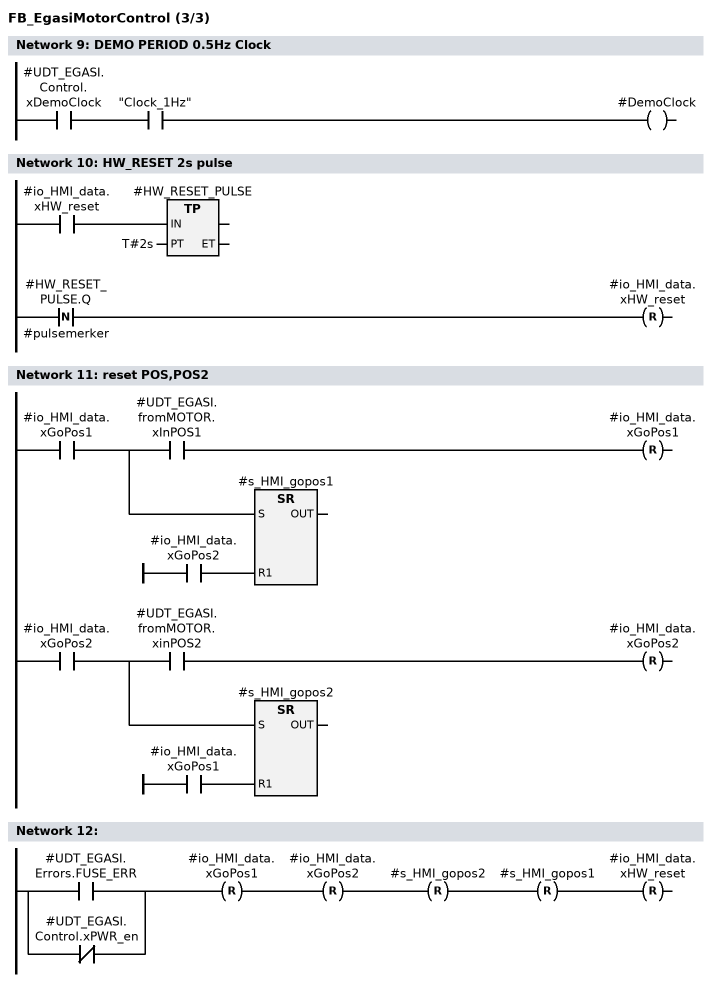
   RUNG wire#powerrail
      Contact( #UDT_EGASI.Control.xDemoClock )
      Contact( "Clock_1Hz" )
      Coil( #DemoClock )
   END_RUNG
   // the same network as SCL:
   #DemoClock := #UDT_EGASI.Control.xDemoClock AND "Clock_1Hz";
END_REGION

REGION Network 10: HW_RESET 2s pulse
   #HW_RESET_PULSE(IN := #io_HMI_data.xHW_reset, PT := T#2s);   // TP
   #_w1 := NOT #HW_RESET_PULSE.Q AND #pulsemerker;   // falling edge of #HW_RESET_PULSE.Q
   #pulsemerker := #HW_RESET_PULSE.Q;
   IF #_w1 THEN #io_HMI_data.xHW_reset := FALSE; END_IF;
END_REGION

REGION Network 11: reset POS,POS2
   RUNG wire#powerrail
      Contact( #io_HMI_data.xGoPos1 )
      wire#w1
      Contact( #UDT_EGASI.fromMOTOR.xInPOS1 )
      R_Coil( #io_HMI_data.xGoPos1 )
   END_RUNG
   RUNG wire#w1
      S_SR(operand := #s_HMI_gopos1, r1 := wire#w2)
   END_RUNG
   RUNG wire#powerrail
      Contact( #io_HMI_data.xGoPos2 )
   END_RUNG wire#w2
   RUNG wire#powerrail
      Contact( #io_HMI_data.xGoPos2 )
      wire#w3
      Contact( #UDT_EGASI.fromMOTOR.xinPOS2 )
      R_Coil( #io_HMI_data.xGoPos2 )
   END_RUNG
   RUNG wire#w3
      S_SR(operand := #s_HMI_gopos2, r1 := wire#w4)
   END_RUNG
   RUNG wire#powerrail
      Contact( #io_HMI_data.xGoPos1 )
   END_RUNG wire#w4
   // the same network as SCL:
   #_w1 := #io_HMI_data.xGoPos1;
   IF #io_HMI_data.xGoPos1 AND #UDT_EGASI.fromMOTOR.xInPOS1 THEN #io_HMI_data.xGoPos1 := FALSE; END_IF;
   IF #_w1 THEN
       #s_HMI_gopos1 := TRUE;   // SR flip-flop
   END_IF;
   IF #io_HMI_data.xGoPos2 THEN #s_HMI_gopos1 := FALSE; END_IF;
   #_w2 := #io_HMI_data.xGoPos2;
   IF #io_HMI_data.xGoPos2 AND #UDT_EGASI.fromMOTOR.xinPOS2 THEN #io_HMI_data.xGoPos2 := FALSE; END_IF;
   IF #_w2 THEN
       #s_HMI_gopos2 := TRUE;   // SR flip-flop
   END_IF;
   IF #io_HMI_data.xGoPos1 THEN #s_HMI_gopos2 := FALSE; END_IF;
END_REGION

REGION Network 12
   RUNG wire#powerrail
      Contact( #UDT_EGASI.Errors.FUSE_ERR )
      wire#w1
      R_Coil( #io_HMI_data.xGoPos1 )
      R_Coil( #io_HMI_data.xGoPos2 )
      R_Coil( #s_HMI_gopos2 )
      R_Coil( #s_HMI_gopos1 )
      R_Coil( #io_HMI_data.xHW_reset )
   END_RUNG
   RUNG wire#powerrail
      I_Contact( #UDT_EGASI.Control.xPWR_en )
   END_RUNG wire#w1
   // the same network as SCL:
   IF #UDT_EGASI.Errors.FUSE_ERR OR NOT #UDT_EGASI.Control.xPWR_en THEN
       #io_HMI_data.xGoPos1 := FALSE;
       #io_HMI_data.xGoPos2 := FALSE;
       #s_HMI_gopos2 := FALSE;
       #s_HMI_gopos1 := FALSE;
       #io_HMI_data.xHW_reset := FALSE;
   END_IF;
END_REGION

REGION Network 13 (SCL)
   #q_rScaledTemperature := ((#i_wRawTempValue/32767.0) * 10.0)/0.04;
   #UDT_EGASI.fromMOTOR.wRawTempValue := #i_wRawTempValue;
   #UDT_EGASI.fromMOTOR.rScaledTempValue := #q_rScaledTemperature;
END_REGION
END_FUNCTION_BLOCK

FUNCTION_BLOCK "FB_Convert16bitToTemperature"   // FB17, LAD
{ S7_Optimized_Access := 'TRUE' }
VERSION : 0.1
   VAR_INPUT
      i_wRawValue : Word;
   END_VAR
   VAR_OUTPUT
      q_uiScaledTemperature : Real;
   END_VAR
BEGIN

REGION Network 2 (SCL)
   #q_uiScaledTemperature := #i_wRawValue/32767.0 * 0.04;
END_REGION
END_FUNCTION_BLOCK

FUNCTION_BLOCK "FB_CYLINDER_CONTROL"   // FB18, LAD
{ S7_Optimized_Access := 'TRUE' }
VERSION : 0.1
   VAR_INPUT
      i_xTrigger : Bool;
      i_udMAXDontProduceFeedCounter : UDInt;
   END_VAR
   VAR_OUTPUT
      q_xM1Output : Bool;
      q_xM2Output : Bool;
      q_xM3Output : Bool;
      q_xM4Output : Bool;
      q_xM5Output : Bool;
   END_VAR
   VAR_IN_OUT
      io_CylinderData : "RRI_izdelki";
      io_LastCylinderData : "RRI_izdelki";
      io_ReceptToMake : "RRI_izdelki";
      io_xChangingPart : Bool;
      io_xuiChangePartCounter : UDInt;
      io_iTrenutniPomik : Int;
      PartNumberForProduction : String;
      LastPartForProduction : String;
   END_VAR
   VAR RETAIN
      markers : Array[0..1] of Bool;
      ChangePartStepCounter : Int;
      iLastPartStVrst : Int;
      iLastPartStCelic : Int;
   END_VAR
   VAR_TEMP   // added for the SCL form of the ladder/FBD networks
      _w1 : Bool;
   END_VAR
BEGIN

REGION Network 1: Povečaj števec za trenutni števec
   // pocečaj trneutni pomik
   // povečaj pomik, če je
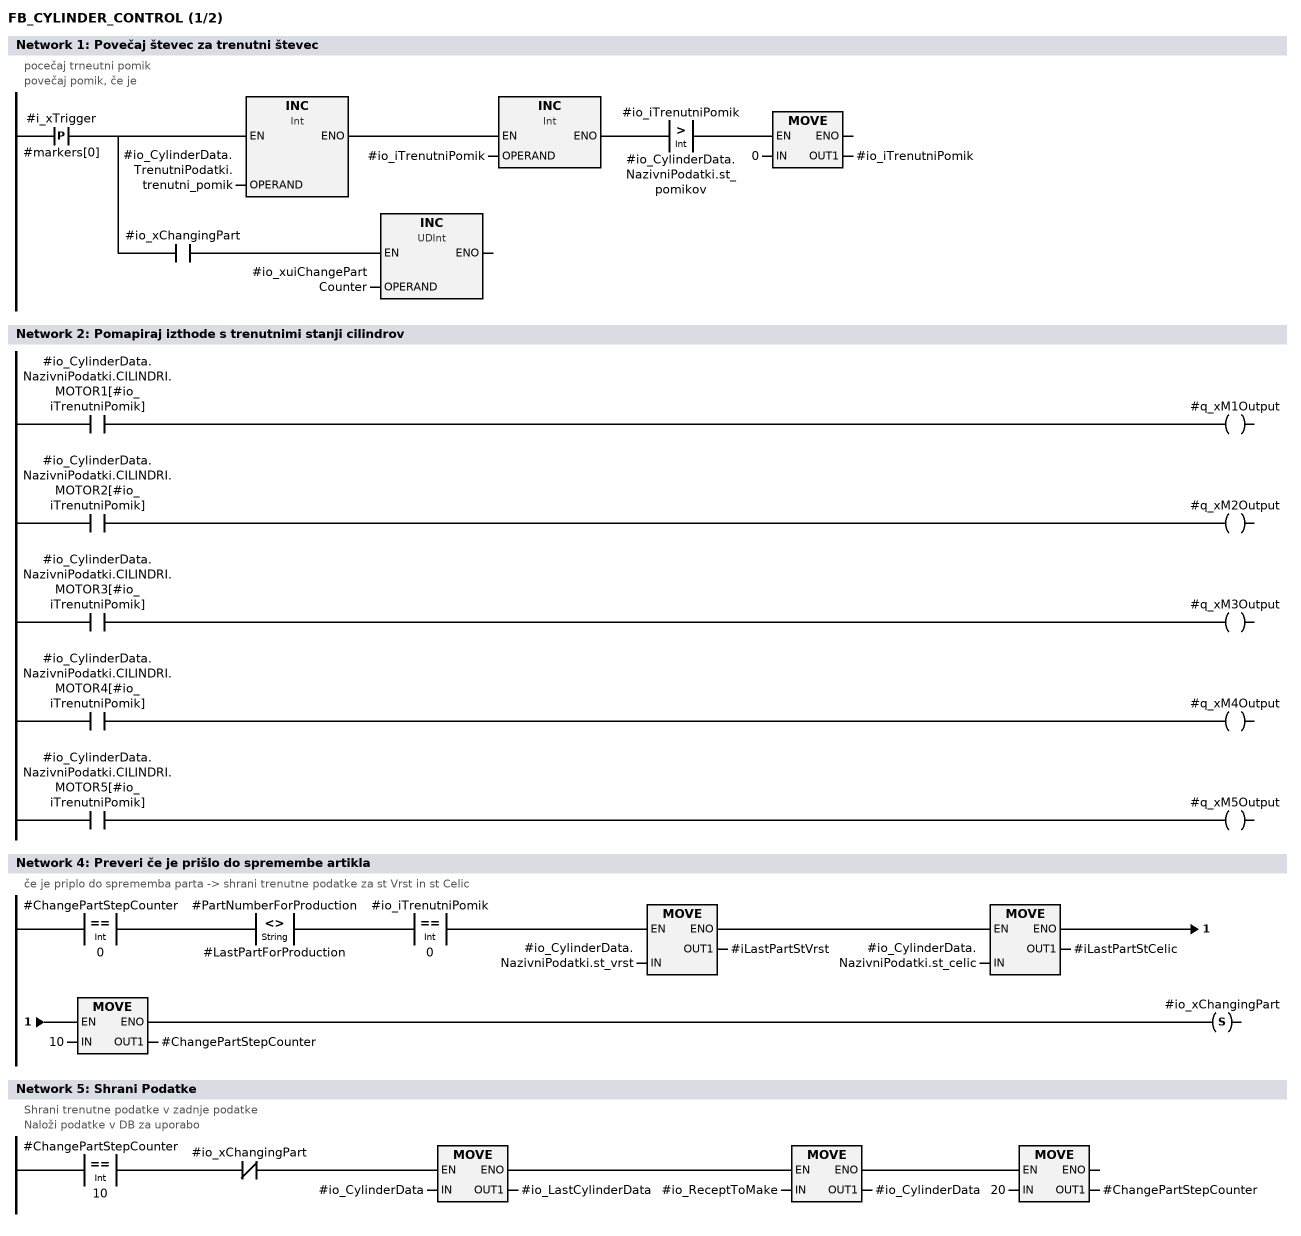
   RUNG wire#powerrail
      P_Contact(operand := #i_xTrigger, bit := #markers[0])
      wire#w1
      { S7_Templates := "DestType := Int" } Inc( #io_CylinderData.TrenutniPodatki.trenutni_pomik )
      { S7_Templates := "DestType := Int" } Inc( #io_iTrenutniPomik )
      { S7_Templates := "SrcType := Int" } GT_Contact(in1 := #io_iTrenutniPomik, in2 := #io_CylinderData.NazivniPodatki.st_pomikov)
      Move(in := 0, out1 => #io_iTrenutniPomik)
   END_RUNG
   RUNG wire#w1
      Contact( #io_xChangingPart )
      { S7_Templates := "DestType := UDInt" } Inc( #io_xuiChangePartCounter )
   END_RUNG
   // the same network as SCL:
   #_w1 := #i_xTrigger AND NOT #markers[0];   // rising edge of #i_xTrigger
   #markers[0] := #i_xTrigger;
   IF #_w1 THEN
       #io_CylinderData.TrenutniPodatki.trenutni_pomik := #io_CylinderData.TrenutniPodatki.trenutni_pomik + 1;
       #io_iTrenutniPomik := #io_iTrenutniPomik + 1;
   END_IF;
   IF #_w1 AND (#io_iTrenutniPomik > #io_CylinderData.NazivniPodatki.st_pomikov) THEN
       #io_iTrenutniPomik := 0;
   END_IF;
   IF #_w1 AND #io_xChangingPart THEN #io_xuiChangePartCounter := #io_xuiChangePartCounter + 1; END_IF;
END_REGION

REGION Network 2: Pomapiraj izthode s trenutnimi stanji cilindrov
   RUNG wire#powerrail
      Contact( #io_CylinderData.NazivniPodatki.CILINDRI.MOTOR1[#io_iTrenutniPomik] )
      Coil( #q_xM1Output )
   END_RUNG
   RUNG wire#powerrail
      Contact( #io_CylinderData.NazivniPodatki.CILINDRI.MOTOR2[#io_iTrenutniPomik] )
      Coil( #q_xM2Output )
   END_RUNG
   RUNG wire#powerrail
      Contact( #io_CylinderData.NazivniPodatki.CILINDRI.MOTOR3[#io_iTrenutniPomik] )
      Coil( #q_xM3Output )
   END_RUNG
   RUNG wire#powerrail
      Contact( #io_CylinderData.NazivniPodatki.CILINDRI.MOTOR4[#io_iTrenutniPomik] )
      Coil( #q_xM4Output )
   END_RUNG
   RUNG wire#powerrail
      Contact( #io_CylinderData.NazivniPodatki.CILINDRI.MOTOR5[#io_iTrenutniPomik] )
      Coil( #q_xM5Output )
   END_RUNG
   // the same network as SCL:
   #q_xM1Output := #io_CylinderData.NazivniPodatki.CILINDRI.MOTOR1[#io_iTrenutniPomik];
   #q_xM2Output := #io_CylinderData.NazivniPodatki.CILINDRI.MOTOR2[#io_iTrenutniPomik];
   #q_xM3Output := #io_CylinderData.NazivniPodatki.CILINDRI.MOTOR3[#io_iTrenutniPomik];
   #q_xM4Output := #io_CylinderData.NazivniPodatki.CILINDRI.MOTOR4[#io_iTrenutniPomik];
   #q_xM5Output := #io_CylinderData.NazivniPodatki.CILINDRI.MOTOR5[#io_iTrenutniPomik];
END_REGION

REGION Network 4: Preveri če je prišlo do spremembe artikla
   // če je priplo do sprememba parta -> shrani trenutne podatke za st Vrst in st Celic
   RUNG wire#powerrail
      { S7_Templates := "SrcType := Int" } EQ_Contact(in1 := #ChangePartStepCounter, in2 := 0)
      { S7_Templates := "SrcType := String" } NE_Contact(in1 := #PartNumberForProduction, in2 := #LastPartForProduction)
      { S7_Templates := "SrcType := Int" } EQ_Contact(in1 := #io_iTrenutniPomik, in2 := 0)
      Move(in := #io_CylinderData.NazivniPodatki.st_vrst, out1 => #iLastPartStVrst)
      Move(in := #io_CylinderData.NazivniPodatki.st_celic, out1 => #iLastPartStCelic)
      Move(in := 10, out1 => #ChangePartStepCounter)
      S_Coil( #io_xChangingPart )
   END_RUNG
   // the same network as SCL:
   IF (#ChangePartStepCounter = 0) AND (#PartNumberForProduction <> #LastPartForProduction) AND (#io_iTrenutniPomik = 0) THEN
       #iLastPartStVrst := #io_CylinderData.NazivniPodatki.st_vrst;
       #iLastPartStCelic := #io_CylinderData.NazivniPodatki.st_celic;
   END_IF;
   #_w1 := (#ChangePartStepCounter = 0) AND (#PartNumberForProduction <> #LastPartForProduction) AND (#io_iTrenutniPomik = 0);
   IF #_w1 THEN
       #ChangePartStepCounter := 10;
       #io_xChangingPart := TRUE;
   END_IF;
END_REGION

REGION Network 5: Shrani Podatke
   // Shrani trenutne podatke v zadnje podatke
   // Naloži podatke v DB za uporabo
   RUNG wire#powerrail
      { S7_Templates := "SrcType := Int" } EQ_Contact(in1 := #ChangePartStepCounter, in2 := 10)
      I_Contact( #io_xChangingPart )
      Move(in := #io_CylinderData, out1 => #io_LastCylinderData)
      Move(in := #io_ReceptToMake, out1 => #io_CylinderData)
      Move(in := 20, out1 => #ChangePartStepCounter)
   END_RUNG
   // the same network as SCL:
   IF (#ChangePartStepCounter = 10) AND NOT #io_xChangingPart THEN
       #io_LastCylinderData := #io_CylinderData;
       #io_CylinderData := #io_ReceptToMake;
       #ChangePartStepCounter := 20;
   END_IF;
END_REGION

REGION Network 6
   // Shrani partnumber
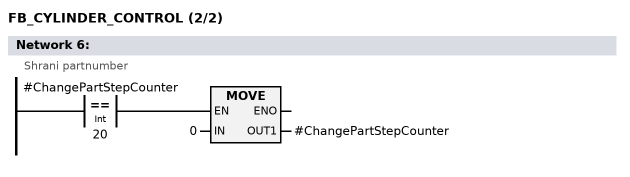
   RUNG wire#powerrail
      { S7_Templates := "SrcType := Int" } EQ_Contact(in1 := #ChangePartStepCounter, in2 := 20)
      Move(in := 0, out1 => #ChangePartStepCounter)
   END_RUNG
   // the same network as SCL:
   IF #ChangePartStepCounter = 20 THEN #ChangePartStepCounter := 0; END_IF;
END_REGION
END_FUNCTION_BLOCK

FUNCTION "FC_INPUT" : Void   // FC1, LAD
{ S7_Optimized_Access := 'TRUE' }
VERSION : 0.1
BEGIN

REGION Network 1: PLC input mapping
   // AKD1 - fault relay - open if error
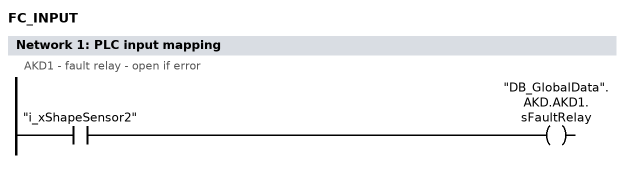
   RUNG wire#powerrail
      Contact( "i_xShapeSensor2" )
      Coil( "DB_GlobalData".AKD.AKD1.sFaultRelay )
   END_RUNG
   // the same network as SCL:
   "DB_GlobalData".AKD.AKD1.sFaultRelay := "i_xShapeSensor2";
END_REGION
END_FUNCTION

FUNCTION "FC_OUTPUT" : Void   // FC2, LAD
{ S7_Optimized_Access := 'TRUE' }
VERSION : 0.1
BEGIN

REGION Network 1: Communication mapping for NodeRed data and DATAFORCOMUNICATIONDB
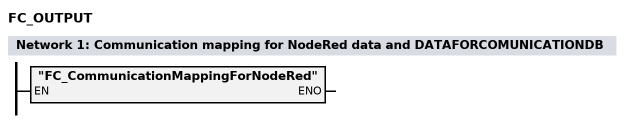
   RUNG wire#powerrail
      "FC_CommunicationMappingForNodeRed"()
   END_RUNG
   // the same network as SCL:
   "FC_CommunicationMappingForNodeRed"();
END_REGION
END_FUNCTION

FUNCTION "FC_LOGIC" : Void   // FC3, LAD
{ S7_Optimized_Access := 'TRUE' }
VERSION : 0.1
BEGIN

REGION Network 1: Convert ThermocuplerData
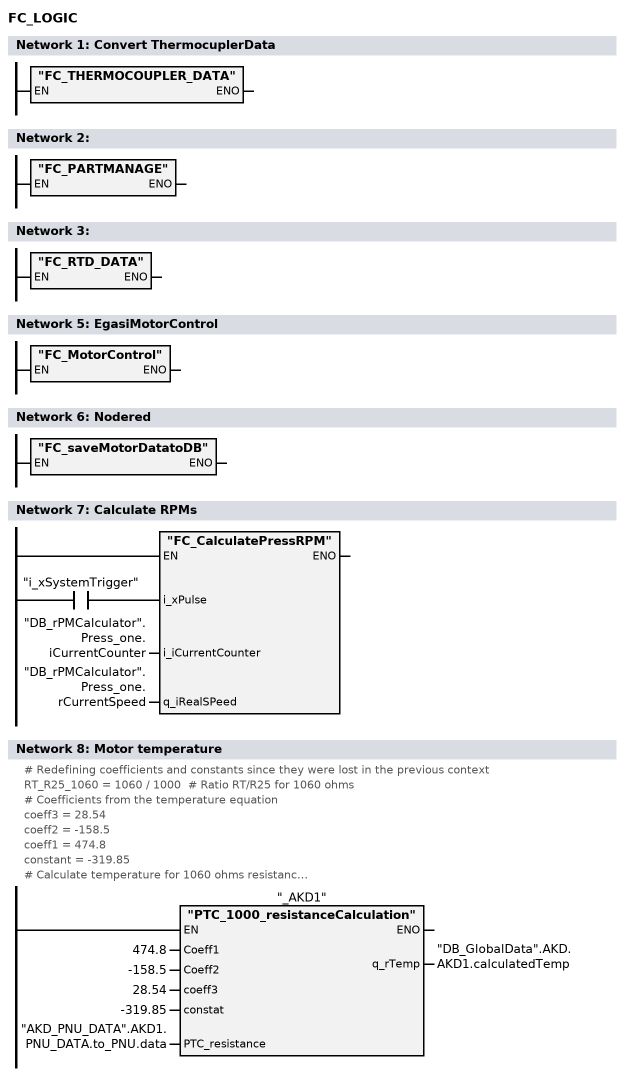
   RUNG wire#powerrail
      "FC_THERMOCOUPLER_DATA"()
   END_RUNG
   // the same network as SCL:
   "FC_THERMOCOUPLER_DATA"();
END_REGION

REGION Network 2
   RUNG wire#powerrail
      "FC_PARTMANAGE"()
   END_RUNG
   // the same network as SCL:
   "FC_PARTMANAGE"();
END_REGION

REGION Network 3
   RUNG wire#powerrail
      "FC_RTD_DATA"()
   END_RUNG
   // the same network as SCL:
   "FC_RTD_DATA"();
END_REGION

REGION Network 4: Kollmorgen Settings
END_REGION

REGION Network 5: EgasiMotorControl
   RUNG wire#powerrail
      "FC_MotorControl"()
   END_RUNG
   // the same network as SCL:
   "FC_MotorControl"();
END_REGION

REGION Network 6: Nodered
   RUNG wire#powerrail
      "FC_saveMotorDatatoDB"()
   END_RUNG
   // the same network as SCL:
   "FC_saveMotorDatatoDB"();
END_REGION

REGION Network 7: Calculate RPMs
   RUNG wire#powerrail
      "FC_CalculatePressRPM"(i_xPulse := wire#w1, i_iCurrentCounter := "DB_rPMCalculator".Press_one.iCurrentCounter, q_iRealSPeed := "DB_rPMCalculator".Press_one.rCurrentSpeed)
   END_RUNG
   RUNG wire#powerrail
      Contact( "i_xSystemTrigger" )
   END_RUNG wire#w1
   // the same network as SCL:
   "FC_CalculatePressRPM"(i_xPulse := "i_xSystemTrigger",
                          i_iCurrentCounter := "DB_rPMCalculator".Press_one.iCurrentCounter,
                          q_iRealSPeed := "DB_rPMCalculator".Press_one.rCurrentSpeed);
END_REGION

REGION Network 8: Motor temperature
   // # Redefining coefficients and constants since they were lost in the previous context
   // RT_R25_1060 = 1060 / 1000  # Ratio RT/R25 for 1060 ohms
   // 
   // # Coefficients from the temperature equation
   // coeff3 = 28.54
   // coeff2 = -158.5
   // coeff1 = 474.8
   // constant = -319.85
   // 
   // # Calculate temperature for 1060 ohms resistance
   // temperature_1060 = (coeff3 * RT_R25_1060**3) + (coeff2 * RT_R25_1060**2) + (coeff1 * RT_R25_1060) + constant
   RUNG wire#powerrail
      "_AKD1"(Coeff1 := 474.8, Coeff2 := -158.5, coeff3 := 28.54, constat := -319.85, PTC_resistance := "AKD_PNU_DATA".AKD1.PNU_DATA.to_PNU.data, q_rTemp => "DB_GlobalData".AKD.AKD1.calculatedTemp)
   END_RUNG
   // the same network as SCL:
   "_AKD1"(Coeff1 := 474.8,   // "PTC_1000_resistanceCalculation"
           Coeff2 := -158.5,
           coeff3 := 28.54,
           constat := -319.85,
           PTC_resistance := "AKD_PNU_DATA".AKD1.PNU_DATA.to_PNU.data,
           q_rTemp => "DB_GlobalData".AKD.AKD1.calculatedTemp);
END_REGION
END_FUNCTION

FUNCTION "FC_THERMOCOUPLER_DATA" : Void   // FC4, LAD
{ S7_Optimized_Access := 'TRUE' }
VERSION : 0.1
BEGIN

REGION Network 1: Temeprature conversion - from Input to GlobalDataBLock
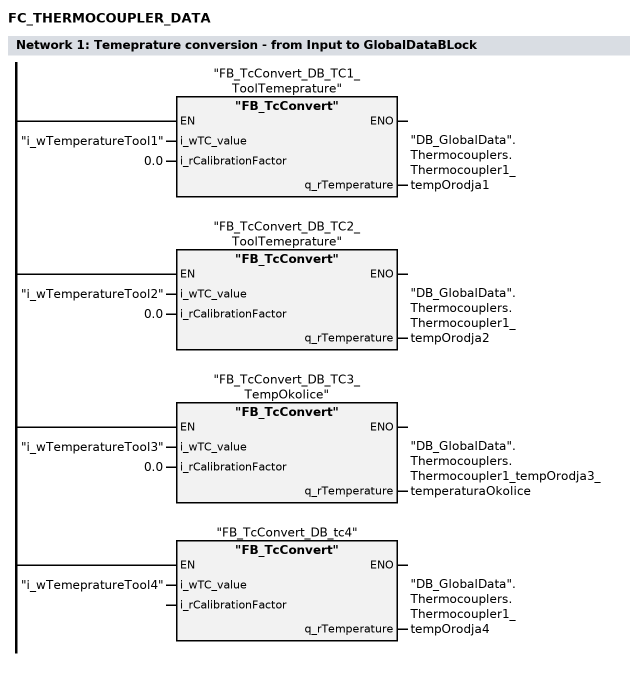
   RUNG wire#powerrail
      "FB_TcConvert_DB_TC1_ToolTemeprature"(i_wTC_value := "i_wTemperatureTool1", i_rCalibrationFactor := 0.0, q_rTemperature => "DB_GlobalData".Thermocouplers.Thermocoupler1_tempOrodja1)
   END_RUNG
   RUNG wire#powerrail
      "FB_TcConvert_DB_TC2_ToolTemeprature"(i_wTC_value := "i_wTemperatureTool2", i_rCalibrationFactor := 0.0, q_rTemperature => "DB_GlobalData".Thermocouplers.Thermocoupler1_tempOrodja2)
   END_RUNG
   RUNG wire#powerrail
      "FB_TcConvert_DB_TC3_TempOkolice"(i_wTC_value := "i_wTemperatureTool3", i_rCalibrationFactor := 0.0, q_rTemperature => "DB_GlobalData".Thermocouplers.Thermocoupler1_tempOrodja3_temperaturaOkolice)
   END_RUNG
   RUNG wire#powerrail
      "FB_TcConvert_DB_tc4"(i_wTC_value := "i_wTemepratureTool4", i_rCalibrationFactor :=, q_rTemperature => "DB_GlobalData".Thermocouplers.Thermocoupler1_tempOrodja4)
   END_RUNG
   // the same network as SCL:
   "FB_TcConvert_DB_TC1_ToolTemeprature"(i_wTC_value := "i_wTemperatureTool1",   // "FB_TcConvert"
                           i_rCalibrationFactor := 0.0,
                           q_rTemperature => "DB_GlobalData".Thermocouplers.Thermocoupler1_tempOrodja1);
   "FB_TcConvert_DB_TC2_ToolTemeprature"(i_wTC_value := "i_wTemperatureTool2",   // "FB_TcConvert"
                           i_rCalibrationFactor := 0.0,
                           q_rTemperature => "DB_GlobalData".Thermocouplers.Thermocoupler1_tempOrodja2);
   "FB_TcConvert_DB_TC3_TempOkolice"(i_wTC_value := "i_wTemperatureTool3",   // "FB_TcConvert"
                           i_rCalibrationFactor := 0.0,
                           q_rTemperature => "DB_GlobalData".Thermocouplers.Thermocoupler1_tempOrodja3_temperaturaOkolice);
   "FB_TcConvert_DB_tc4"(i_wTC_value := "i_wTemepratureTool4",   // "FB_TcConvert"
                         q_rTemperature => "DB_GlobalData".Thermocouplers.Thermocoupler1_tempOrodja4);
END_REGION
END_FUNCTION

FUNCTION "FC_CommunicationMappingForNodeRed" : Void   // FC5, LAD
{ S7_Optimized_Access := 'TRUE' }
VERSION : 0.1
   VAR_TEMP   // added for the SCL form of the ladder/FBD networks
      _w1 : Bool;
   END_VAR
BEGIN

REGION Network 1: Move data from GlobalData to DB for NodeRedCommunication
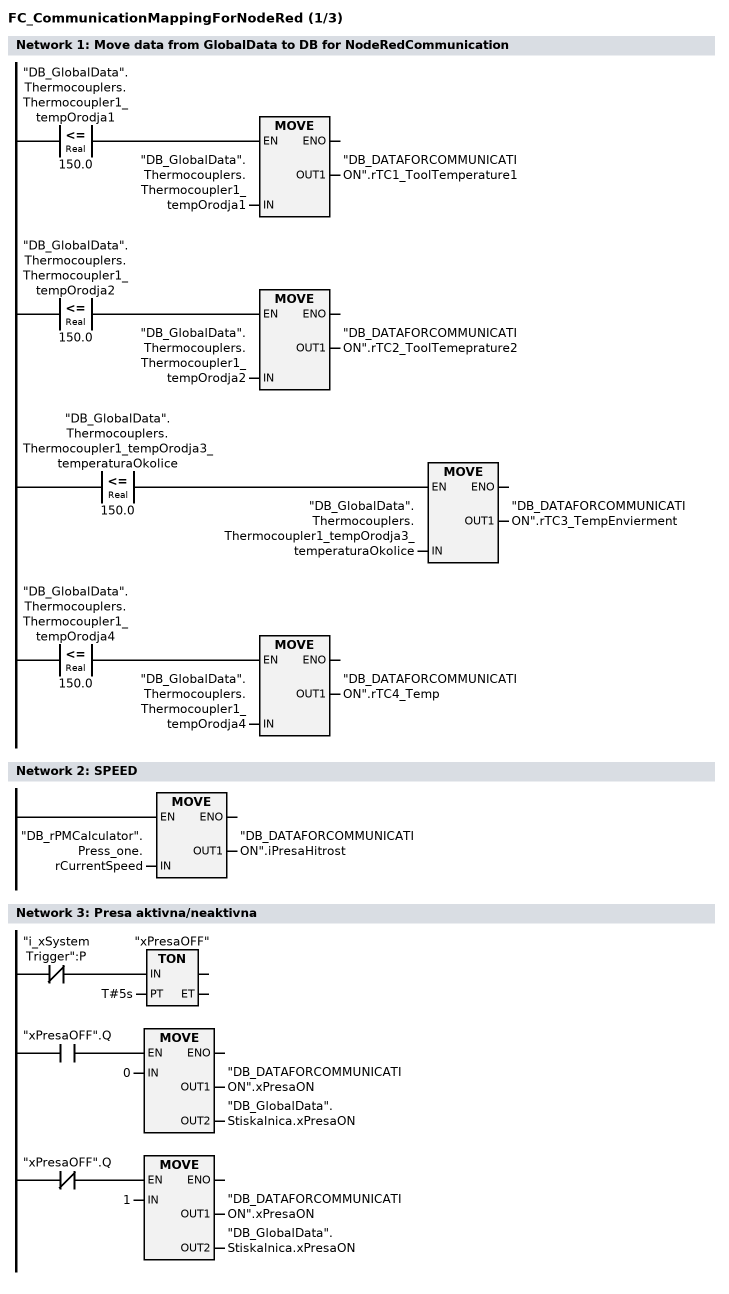
   RUNG wire#powerrail
      { S7_Templates := "SrcType := Real" } LE_Contact(in1 := "DB_GlobalData".Thermocouplers.Thermocoupler1_tempOrodja1, in2 := 150.0)
      Move(in := "DB_GlobalData".Thermocouplers.Thermocoupler1_tempOrodja1, out1 => "DB_DATAFORCOMMUNICATION".rTC1_ToolTemperature1)
   END_RUNG
   RUNG wire#powerrail
      { S7_Templates := "SrcType := Real" } LE_Contact(in1 := "DB_GlobalData".Thermocouplers.Thermocoupler1_tempOrodja2, in2 := 150.0)
      Move(in := "DB_GlobalData".Thermocouplers.Thermocoupler1_tempOrodja2, out1 => "DB_DATAFORCOMMUNICATION".rTC2_ToolTemeprature2)
   END_RUNG
   RUNG wire#powerrail
      { S7_Templates := "SrcType := Real" } LE_Contact(in1 := "DB_GlobalData".Thermocouplers.Thermocoupler1_tempOrodja3_temperaturaOkolice, in2 := 150.0)
      Move(in := "DB_GlobalData".Thermocouplers.Thermocoupler1_tempOrodja3_temperaturaOkolice, out1 => "DB_DATAFORCOMMUNICATION".rTC3_TempEnvierment)
   END_RUNG
   RUNG wire#powerrail
      { S7_Templates := "SrcType := Real" } LE_Contact(in1 := "DB_GlobalData".Thermocouplers.Thermocoupler1_tempOrodja4, in2 := 150.0)
      Move(in := "DB_GlobalData".Thermocouplers.Thermocoupler1_tempOrodja4, out1 => "DB_DATAFORCOMMUNICATION".rTC4_Temp)
   END_RUNG
   // the same network as SCL:
   IF "DB_GlobalData".Thermocouplers.Thermocoupler1_tempOrodja1 <= 150.0 THEN
       "DB_DATAFORCOMMUNICATION".rTC1_ToolTemperature1 := "DB_GlobalData".Thermocouplers.Thermocoupler1_tempOrodja1;
   END_IF;
   IF "DB_GlobalData".Thermocouplers.Thermocoupler1_tempOrodja2 <= 150.0 THEN
       "DB_DATAFORCOMMUNICATION".rTC2_ToolTemeprature2 := "DB_GlobalData".Thermocouplers.Thermocoupler1_tempOrodja2;
   END_IF;
   IF "DB_GlobalData".Thermocouplers.Thermocoupler1_tempOrodja3_temperaturaOkolice <= 150.0 THEN
       "DB_DATAFORCOMMUNICATION".rTC3_TempEnvierment := "DB_GlobalData".Thermocouplers.Thermocoupler1_tempOrodja3_temperaturaOkolice;
   END_IF;
   IF "DB_GlobalData".Thermocouplers.Thermocoupler1_tempOrodja4 <= 150.0 THEN
       "DB_DATAFORCOMMUNICATION".rTC4_Temp := "DB_GlobalData".Thermocouplers.Thermocoupler1_tempOrodja4;
   END_IF;
END_REGION

REGION Network 2: SPEED
   RUNG wire#powerrail
      Move(in := "DB_rPMCalculator".Press_one.rCurrentSpeed, out1 => "DB_DATAFORCOMMUNICATION".iPresaHitrost)
   END_RUNG
   // the same network as SCL:
   "DB_DATAFORCOMMUNICATION".iPresaHitrost := "DB_rPMCalculator".Press_one.rCurrentSpeed;
END_REGION

REGION Network 3: Presa aktivna/neaktivna
   "xPresaOFF".TON(IN := NOT "i_xSystemTrigger":P, PT := T#5s);
   IF "xPresaOFF".Q THEN
       "DB_DATAFORCOMMUNICATION".xPresaON := 0;
       "DB_GlobalData".Stiskalnica.xPresaON := 0;
   END_IF;
   IF NOT "xPresaOFF".Q THEN
       "DB_DATAFORCOMMUNICATION".xPresaON := 1;
       "DB_GlobalData".Stiskalnica.xPresaON := 1;
   END_IF;
END_REGION

REGION Network 4: Stevec preklopov
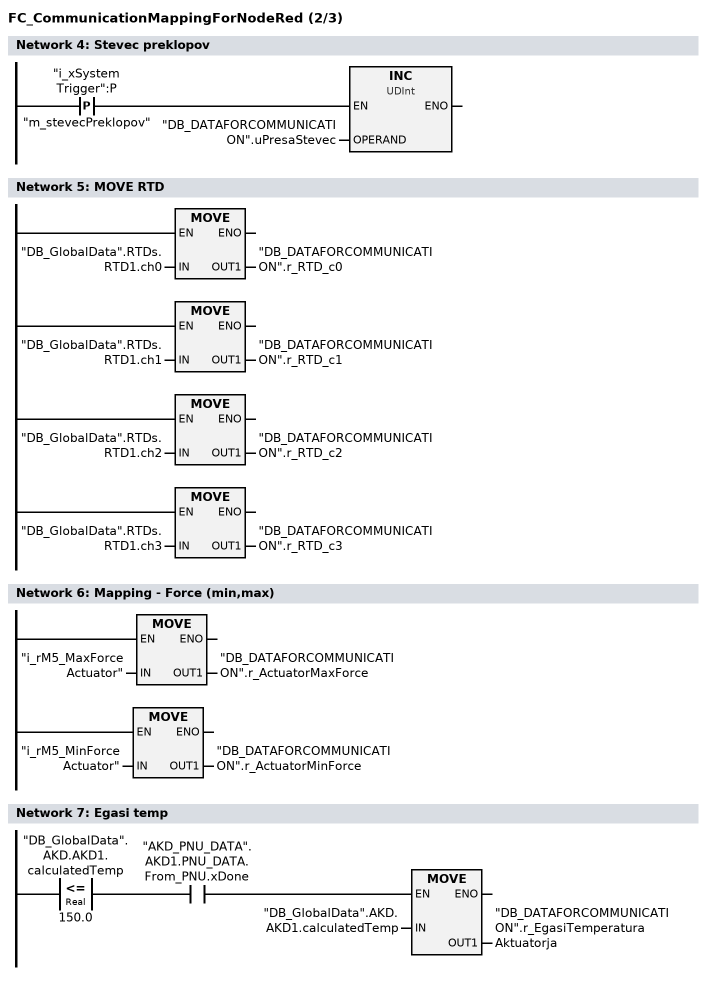
   RUNG wire#powerrail
      P_Contact(operand := "i_xSystemTrigger":P, bit := "m_stevecPreklopov")
      { S7_Templates := "DestType := UDInt" } Inc( "DB_DATAFORCOMMUNICATION".uPresaStevec )
   END_RUNG
   // the same network as SCL:
   #_w1 := "i_xSystemTrigger":P AND NOT "m_stevecPreklopov";   // rising edge of "i_xSystemTrigger":P
   "m_stevecPreklopov" := "i_xSystemTrigger":P;
   IF #_w1 THEN "DB_DATAFORCOMMUNICATION".uPresaStevec := "DB_DATAFORCOMMUNICATION".uPresaStevec + 1; END_IF;
END_REGION

REGION Network 5: MOVE RTD
   RUNG wire#powerrail
      Move(in := "DB_GlobalData".RTDs.RTD1.ch0, out1 => "DB_DATAFORCOMMUNICATION".r_RTD_c0)
   END_RUNG
   RUNG wire#powerrail
      Move(in := "DB_GlobalData".RTDs.RTD1.ch1, out1 => "DB_DATAFORCOMMUNICATION".r_RTD_c1)
   END_RUNG
   RUNG wire#powerrail
      Move(in := "DB_GlobalData".RTDs.RTD1.ch2, out1 => "DB_DATAFORCOMMUNICATION".r_RTD_c2)
   END_RUNG
   RUNG wire#powerrail
      Move(in := "DB_GlobalData".RTDs.RTD1.ch3, out1 => "DB_DATAFORCOMMUNICATION".r_RTD_c3)
   END_RUNG
   // the same network as SCL:
   "DB_DATAFORCOMMUNICATION".r_RTD_c0 := "DB_GlobalData".RTDs.RTD1.ch0;
   "DB_DATAFORCOMMUNICATION".r_RTD_c1 := "DB_GlobalData".RTDs.RTD1.ch1;
   "DB_DATAFORCOMMUNICATION".r_RTD_c2 := "DB_GlobalData".RTDs.RTD1.ch2;
   "DB_DATAFORCOMMUNICATION".r_RTD_c3 := "DB_GlobalData".RTDs.RTD1.ch3;
END_REGION

REGION Network 6: Mapping - Force (min,max)
   RUNG wire#powerrail
      Move(in := "i_rM5_MaxForceActuator", out1 => "DB_DATAFORCOMMUNICATION".r_ActuatorMaxForce)
   END_RUNG
   RUNG wire#powerrail
      Move(in := "i_rM5_MinForceActuator", out1 => "DB_DATAFORCOMMUNICATION".r_ActuatorMinForce)
   END_RUNG
   // the same network as SCL:
   "DB_DATAFORCOMMUNICATION".r_ActuatorMaxForce := "i_rM5_MaxForceActuator";
   "DB_DATAFORCOMMUNICATION".r_ActuatorMinForce := "i_rM5_MinForceActuator";
END_REGION

REGION Network 7: Egasi temp
   RUNG wire#powerrail
      { S7_Templates := "SrcType := Real" } LE_Contact(in1 := "DB_GlobalData".AKD.AKD1.calculatedTemp, in2 := 150.0)
      Contact( "AKD_PNU_DATA".AKD1.PNU_DATA.From_PNU.xDone )
      Move(in := "DB_GlobalData".AKD.AKD1.calculatedTemp, out1 => "DB_DATAFORCOMMUNICATION".r_EgasiTemperaturaAktuatorja)
   END_RUNG
   // the same network as SCL:
   IF ("DB_GlobalData".AKD.AKD1.calculatedTemp <= 150.0) AND "AKD_PNU_DATA".AKD1.PNU_DATA.From_PNU.xDone THEN
       "DB_DATAFORCOMMUNICATION".r_EgasiTemperaturaAktuatorja := "DB_GlobalData".AKD.AKD1.calculatedTemp;
   END_IF;
END_REGION

REGION Network 8: EGASI MOTOR
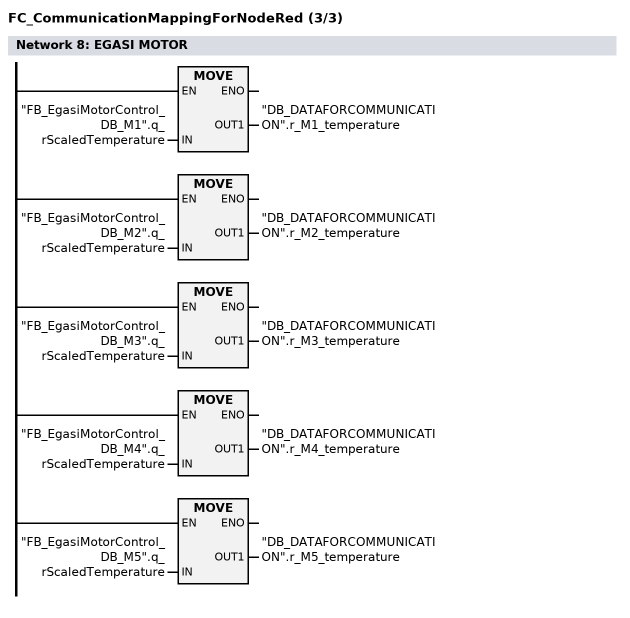
   RUNG wire#powerrail
      Move(in := "FB_EgasiMotorControl_DB_M1".q_rScaledTemperature, out1 => "DB_DATAFORCOMMUNICATION".r_M1_temperature)
   END_RUNG
   RUNG wire#powerrail
      Move(in := "FB_EgasiMotorControl_DB_M2".q_rScaledTemperature, out1 => "DB_DATAFORCOMMUNICATION".r_M2_temperature)
   END_RUNG
   RUNG wire#powerrail
      Move(in := "FB_EgasiMotorControl_DB_M3".q_rScaledTemperature, out1 => "DB_DATAFORCOMMUNICATION".r_M3_temperature)
   END_RUNG
   RUNG wire#powerrail
      Move(in := "FB_EgasiMotorControl_DB_M4".q_rScaledTemperature, out1 => "DB_DATAFORCOMMUNICATION".r_M4_temperature)
   END_RUNG
   RUNG wire#powerrail
      Move(in := "FB_EgasiMotorControl_DB_M5".q_rScaledTemperature, out1 => "DB_DATAFORCOMMUNICATION".r_M5_temperature)
   END_RUNG
   // the same network as SCL:
   "DB_DATAFORCOMMUNICATION".r_M1_temperature := "FB_EgasiMotorControl_DB_M1".q_rScaledTemperature;
   "DB_DATAFORCOMMUNICATION".r_M2_temperature := "FB_EgasiMotorControl_DB_M2".q_rScaledTemperature;
   "DB_DATAFORCOMMUNICATION".r_M3_temperature := "FB_EgasiMotorControl_DB_M3".q_rScaledTemperature;
   "DB_DATAFORCOMMUNICATION".r_M4_temperature := "FB_EgasiMotorControl_DB_M4".q_rScaledTemperature;
   "DB_DATAFORCOMMUNICATION".r_M5_temperature := "FB_EgasiMotorControl_DB_M5".q_rScaledTemperature;
END_REGION
END_FUNCTION

FUNCTION "FC_AKD_KOLLMORGEN" : Void   // FC6, LAD
{ S7_Optimized_Access := 'TRUE' }
VERSION : 0.1
   VAR_TEMP   // added for the SCL form of the ladder/FBD networks
      _w1 : Bool;
      _w2 : Bool;
   END_VAR
BEGIN

REGION Network 1: AKD1
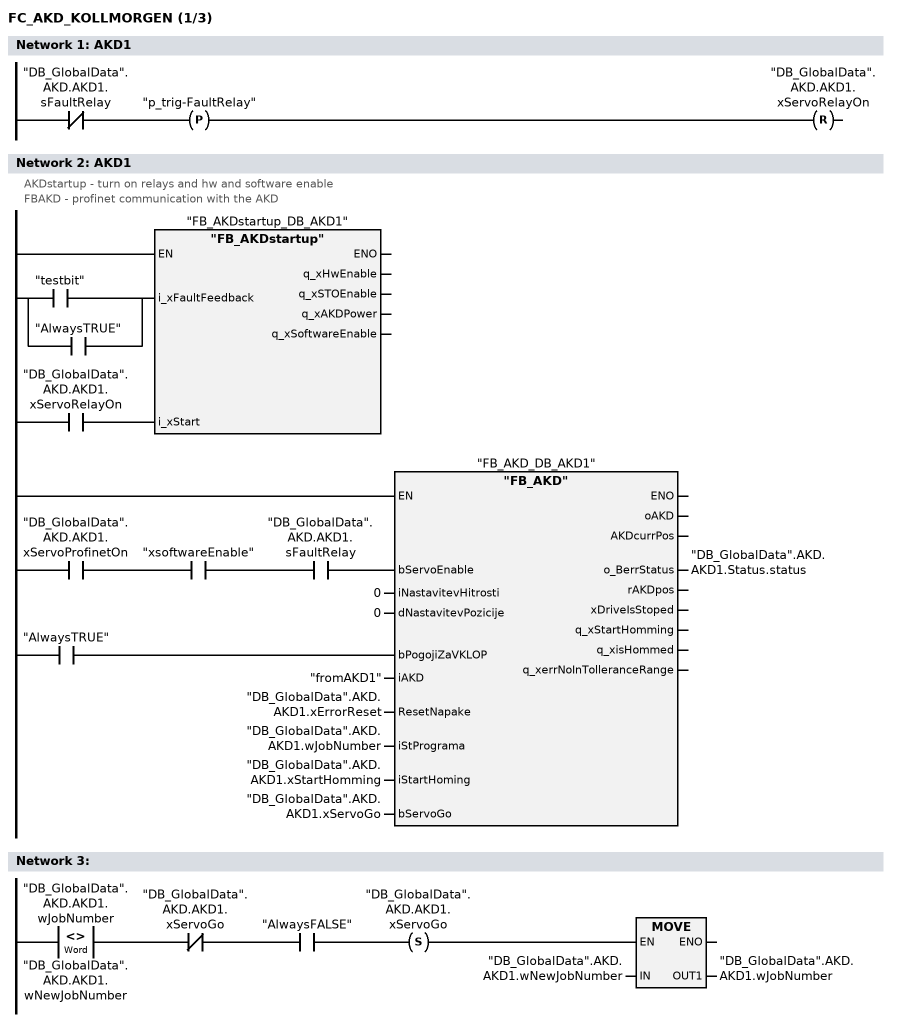
   RUNG wire#powerrail
      I_Contact( "DB_GlobalData".AKD.AKD1.sFaultRelay )
      P_Trig( "p_trig-FaultRelay" )
      R_Coil( "DB_GlobalData".AKD.AKD1.xServoRelayOn )
   END_RUNG
   // the same network as SCL:
   #_w1 := NOT "DB_GlobalData".AKD.AKD1.sFaultRelay AND NOT "p_trig-FaultRelay";   // rising edge
   "p_trig-FaultRelay" := NOT "DB_GlobalData".AKD.AKD1.sFaultRelay;
   IF #_w1 THEN "DB_GlobalData".AKD.AKD1.xServoRelayOn := FALSE; END_IF;
END_REGION

REGION Network 2: AKD1
   // AKDstartup - turn on relays and hw and software enable
   // FBAKD - profinet communication with the AKD
   RUNG wire#powerrail
      "FB_AKDstartup_DB_AKD1"(i_xFaultFeedback := wire#w1, i_xStart := wire#w2, q_xHwEnable =>, q_xSTOEnable =>, q_xAKDPower =>, q_xSoftwareEnable =>)
   END_RUNG
   RUNG wire#powerrail
      Contact( "testbit" )
   END_RUNG wire#w1
   RUNG wire#powerrail
      Contact( "AlwaysTRUE" )
   END_RUNG wire#w1
   RUNG wire#powerrail
      Contact( "DB_GlobalData".AKD.AKD1.xServoRelayOn )
   END_RUNG wire#w2
   RUNG wire#powerrail
      "FB_AKD_DB_AKD1"(bServoEnable := wire#w3, bPogojiZaVKLOP := wire#w4, iNastavitevHitrosti := 0, dNastavitevPozicije := 0, iAKD := "fromAKD1", ResetNapake := "DB_GlobalData".AKD.AKD1.xErrorReset, iStPrograma := "DB_GlobalData".AKD.AKD1.wJobNumber, iStartHoming := "DB_GlobalData".AKD.AKD1.xStartHomming, bServoGo := "DB_GlobalData".AKD.AKD1.xServoGo, oAKD =>, AKDcurrPos =>, o_BerrStatus => "DB_GlobalData".AKD.AKD1.Status.status, rAKDpos =>, xDriveIsStoped =>, q_xStartHomming =>, q_xisHommed =>, q_xerrNoInTolleranceRange =>)
   END_RUNG
   RUNG wire#powerrail
      Contact( "DB_GlobalData".AKD.AKD1.xServoProfinetOn )
      Contact( "xsoftwareEnable" )
      Contact( "DB_GlobalData".AKD.AKD1.sFaultRelay )
   END_RUNG wire#w3
   RUNG wire#powerrail
      Contact( "AlwaysTRUE" )
   END_RUNG wire#w4
   // the same network as SCL:
   "FB_AKDstartup_DB_AKD1"(i_xFaultFeedback := "testbit" OR "AlwaysTRUE",   // "FB_AKDstartup"
                           i_xStart := "DB_GlobalData".AKD.AKD1.xServoRelayOn);
   "FB_AKD_DB_AKD1"(bServoEnable := "DB_GlobalData".AKD.AKD1.xServoProfinetOn AND "xsoftwareEnable" AND "DB_GlobalData".AKD.AKD1.sFaultRelay,   // "FB_AKD"
                    iNastavitevHitrosti := 0,
                    dNastavitevPozicije := 0,
                    bPogojiZaVKLOP := "AlwaysTRUE",
                    iAKD := "fromAKD1",
                    ResetNapake := "DB_GlobalData".AKD.AKD1.xErrorReset,
                    iStPrograma := "DB_GlobalData".AKD.AKD1.wJobNumber,
                    iStartHoming := "DB_GlobalData".AKD.AKD1.xStartHomming,
                    bServoGo := "DB_GlobalData".AKD.AKD1.xServoGo,
                    o_BerrStatus => "DB_GlobalData".AKD.AKD1.Status.status);
END_REGION

REGION Network 3
   RUNG wire#powerrail
      { S7_Templates := "SrcType := Word" } NE_Contact(in1 := "DB_GlobalData".AKD.AKD1.wJobNumber, in2 := "DB_GlobalData".AKD.AKD1.wNewJobNumber)
      I_Contact( "DB_GlobalData".AKD.AKD1.xServoGo )
      Contact( "AlwaysFALSE" )
      S_Coil( "DB_GlobalData".AKD.AKD1.xServoGo )
      Move(in := "DB_GlobalData".AKD.AKD1.wNewJobNumber, out1 => "DB_GlobalData".AKD.AKD1.wJobNumber)
   END_RUNG
   // the same network as SCL:
   #_w1 := ("DB_GlobalData".AKD.AKD1.wJobNumber <> "DB_GlobalData".AKD.AKD1.wNewJobNumber) AND NOT "DB_GlobalData".AKD.AKD1.xServoGo AND "AlwaysFALSE";
   IF #_w1 THEN
       "DB_GlobalData".AKD.AKD1.xServoGo := TRUE;
       "DB_GlobalData".AKD.AKD1.wJobNumber := "DB_GlobalData".AKD.AKD1.wNewJobNumber;
   END_IF;
END_REGION

REGION Network 4: DEMO mode - JOB 0 - 1
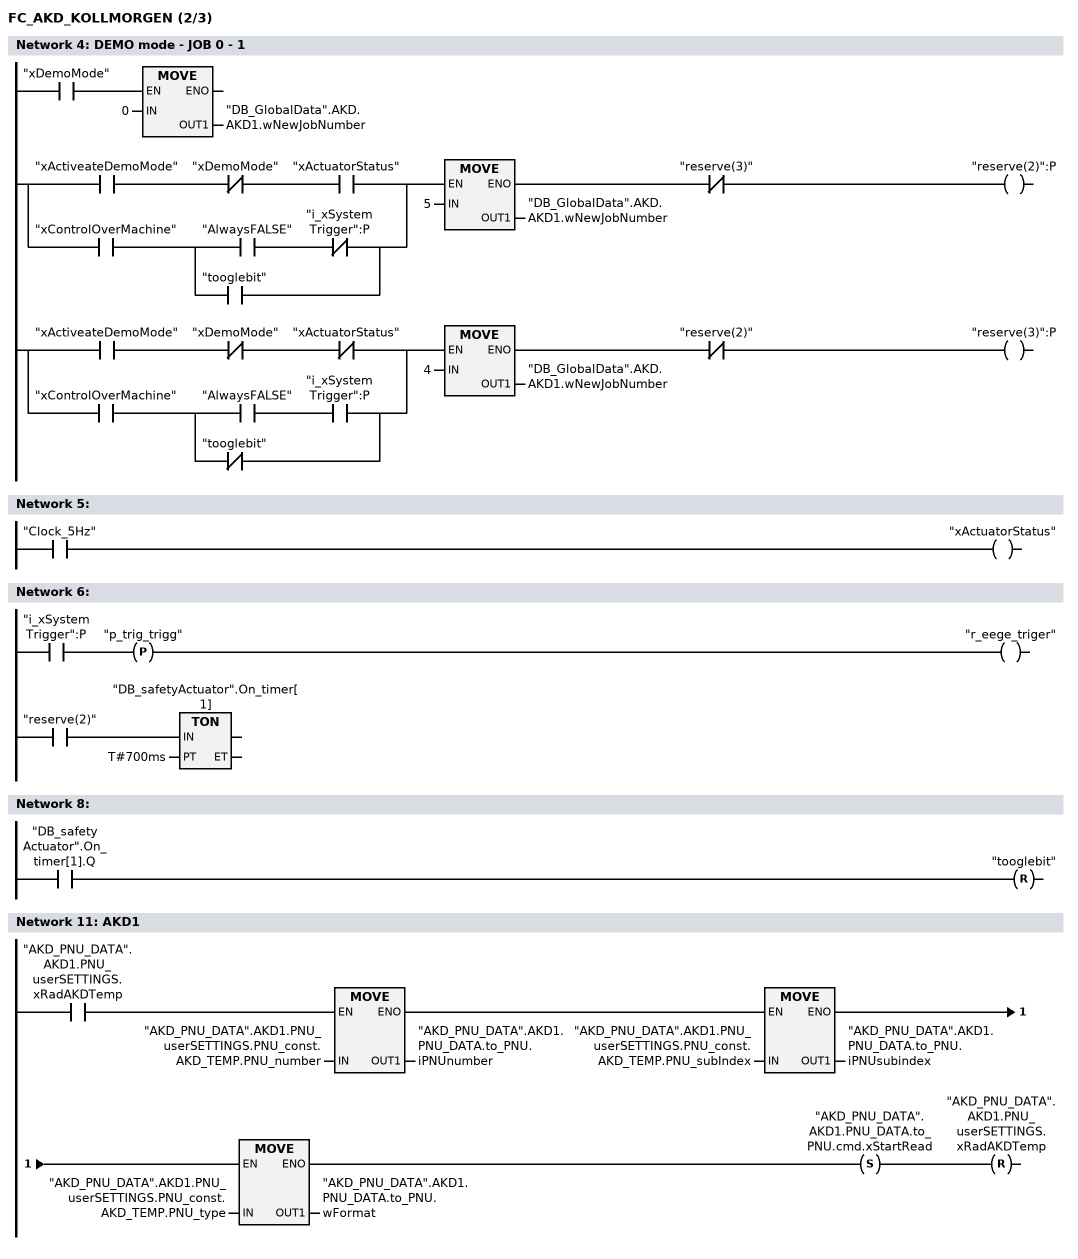
   RUNG wire#powerrail
      Contact( "xDemoMode" )
      Move(in := 0, out1 => "DB_GlobalData".AKD.AKD1.wNewJobNumber)
   END_RUNG
   RUNG wire#powerrail
      Contact( "xActiveateDemoMode" )
      I_Contact( "xDemoMode" )
      Contact( "xActuatorStatus" )
      wire#w1
      Move(in := 5, out1 => "DB_GlobalData".AKD.AKD1.wNewJobNumber)
      I_Contact( "reserve(3)" )
      Coil( "reserve(2)":P )
   END_RUNG
   RUNG wire#powerrail
      Contact( "xControlOverMachine" )
      wire#w2
      Contact( "AlwaysFALSE" )
      I_Contact( "i_xSystemTrigger":P )
   END_RUNG wire#w1
   RUNG wire#w2
      Contact( "tooglebit" )
   END_RUNG wire#w1
   RUNG wire#powerrail
      Contact( "xActiveateDemoMode" )
      I_Contact( "xDemoMode" )
      I_Contact( "xActuatorStatus" )
      wire#w3
      Move(in := 4, out1 => "DB_GlobalData".AKD.AKD1.wNewJobNumber)
      I_Contact( "reserve(2)" )
      Coil( "reserve(3)":P )
   END_RUNG
   RUNG wire#powerrail
      Contact( "xControlOverMachine" )
      wire#w4
      Contact( "AlwaysFALSE" )
      Contact( "i_xSystemTrigger":P )
   END_RUNG wire#w3
   RUNG wire#w4
      I_Contact( "tooglebit" )
   END_RUNG wire#w3
   // the same network as SCL:
   IF "xDemoMode" THEN "DB_GlobalData".AKD.AKD1.wNewJobNumber := 0; END_IF;
   #_w1 := ("xActiveateDemoMode" AND NOT "xDemoMode" AND "xActuatorStatus") OR ("xControlOverMachine" AND (("AlwaysFALSE" AND NOT "i_xSystemTrigger":P) OR "tooglebit"));
   IF #_w1 THEN "DB_GlobalData".AKD.AKD1.wNewJobNumber := 5; END_IF;
   "reserve(2)":P := #_w1 AND NOT "reserve(3)";
   #_w2 := ("xActiveateDemoMode" AND NOT "xDemoMode" AND NOT "xActuatorStatus") OR ("xControlOverMachine" AND (("AlwaysFALSE" AND "i_xSystemTrigger":P) OR NOT "tooglebit"));